
screen "33_Mode_Station_3" 800x480
   Button "Button_5" at 299,208 size 88x48; TextOff 'Stop / AUTO'
      on Press: SetTag("DB_HMI_ARG1_Seq1_Cmd_Auto(2)", 1)
      on Release: SetTag("DB_HMI_ARG1_Seq1_Cmd_Auto(2)", 0)
   Button "Button_6" at 405,208 size 88x48; TextOff 'Reset / MAN'
      on Press: SetTag("DB_HMI_ARG1_Seq1_Cmd_Man(2)", 1)
      on Release: SetTag("DB_HMI_ARG1_Seq1_Cmd_Man(2)", 0)
   Button "Button_1" at 177,283 size 440x40; TextOn 'CLOSE / SCHLIESSEN'; TextOff 'CLOSE / SCHLIESSEN'
      on Click: function_efd93a16()
      Appearance <- "ButtonDown"
   TextField "txtTitleBar" at 16,8 size 495x32; Text 'Operating Mode / Betriebsmodus'
   TextField "txtParameter7_3" at 193,122 size 163x24; Text 'Current Mode / Aktueller Modus'
   TextField "Auto" at 193,149 size 37x20; Text 'Auto'
      Visibility <- "DB_HMI_ARG1_Seq1_Status_Auto(2)"
   TextField "Manual" at 193,148 size 32x20; Text 'Man'
      Visibility <- "DB_HMI_ARG1_Seq1_Status_Man(2)"

screen "34_Mode_Station_4" 800x480
   Button "Button_5" at 299,208 size 88x48; TextOff 'Stop / AUTO'
      on Press: SetTag("DB_HMI_ARG1_Seq1_Cmd_Auto(3)", 1)
      on Release: SetTag("DB_HMI_ARG1_Seq1_Cmd_Auto(3)", 0)
   Button "Button_6" at 405,208 size 88x48; TextOff 'Reset / MAN'
      on Press: SetTag("DB_HMI_ARG1_Seq1_Cmd_Man(3)", 1)
      on Release: SetTag("DB_HMI_ARG1_Seq1_Cmd_Man(3)", 0)
   Button "Button_1" at 177,283 size 440x40; TextOn 'CLOSE / SCHLIESSEN'; TextOff 'CLOSE / SCHLIESSEN'
      on Click: function_efd93a16()
      Appearance <- "ButtonDown"
   TextField "txtTitleBar" at 16,8 size 495x32; Text 'Operating Mode / Betriebsmodus'
   TextField "txtParameter7_3" at 193,122 size 163x24; Text 'Current Mode / Aktueller Modus'
   TextField "Auto" at 193,149 size 37x20; Text 'Auto'
      Visibility <- "DB_HMI_ARG1_Seq1_Status_Auto(3)"
   TextField "Manual" at 193,148 size 32x20; Text 'Man'
      Visibility <- "DB_HMI_ARG1_Seq1_Status_Man(3)"

screen "35_Mode_Station_5" 800x480
   Button "Button_5" at 299,208 size 88x48; TextOff 'Stop / AUTO'
      on Press: SetTag("DB_HMI_ARG1_Seq1_Cmd_Auto(4)", 1)
      on Release: SetTag("DB_HMI_ARG1_Seq1_Cmd_Auto(4)", 0)
   Button "Button_6" at 405,208 size 88x48; TextOff 'Reset / MAN'
      on Press: SetTag("DB_HMI_ARG1_Seq1_Cmd_Man(4)", 1)
      on Release: SetTag("DB_HMI_ARG1_Seq1_Cmd_Man(4)", 0)
   Button "Button_1" at 177,283 size 440x40; TextOn 'CLOSE / SCHLIESSEN'; TextOff 'CLOSE / SCHLIESSEN'
      on Click: function_efd93a16()
      Appearance <- "ButtonDown"
   TextField "txtTitleBar" at 16,8 size 495x32; Text 'Operating Mode / Betriebsmodus'
   TextField "txtParameter7_3" at 193,122 size 163x24; Text 'Current Mode / Aktueller Modus'
   TextField "Auto" at 193,149 size 37x20; Text 'Auto'
      Visibility <- "DB_HMI_ARG1_Seq1_Status_Auto(4)"
   TextField "Manual" at 193,148 size 32x20; Text 'Man'
      Visibility <- "DB_HMI_ARG1_Seq1_Status_Man(4)"

screen "40_SimValues_1" 800x480, template "31_SimValues_1"
   GraphicView "gfxDarkBackground" at 0,0 size 800x480; Picture "PopUpBackground"
      Visibility <- "PopUpBackground"
   TextField "txtParameter1_2" at 246,136 size 42x25; Text 'Step 2 / Parameter 1'
   TextField "txtParameter1_3" at 316,136 size 102x25; Text 'Step 3 / Parameter 1'
   TextField "txtParameter1_4" at 386,136 size 102x25; Text 'Step 4 / Parameter 1'
   TextField "txtParameter1_5" at 456,136 size 102x25; Text 'Step 5 / Parameter 1'
   TextField "txtParameter1_6" at 526,136 size 102x25; Text 'Step 6 / Parameter 1'
   TextField "txtParameter1_8" at 596,136 size 102x25; Text 'Step 7 / Parameter 1'
   TextField "txtParameter1_9" at 666,136 size 102x25; Text 'Step 8 / Parameter 1'
   TextField "txtParameter1_10" at 176,136 size 45x25; Text 'Step 1 / Parameter 1'
   TextField "txtParameter1_11" at 736,136 size 46x25; Text 'Step 9 / Parameter 1'
   TextField "txtParameter1_1" at 104,136 size 45x25; Text 'Branch / Parameter 1'
   TextField "txtParameter1_7" at 32,136 size 45x25; Text 'Car / Parameter 1'
   GraphicView "Graphic view_1" at 33,184 size 40x40; Picture "Car_Red"
   GraphicView "Graphic view_3" at 33,249 size 40x40; Picture "Car_Green"
   GraphicView "Graphic view_4" at 33,308 size 40x40; Picture "Car_Blue_1"
   TextField "Text field_3" at 121,191 size 15x23; Text '1'
      Visibility <- "InScreenTabState"
   TextField "Text field_1" at 121,256 size 15x23; Text '2'
      Visibility <- "InScreenTabState"
   TextField "Text field_2" at 121,321 size 15x23; Text '2'
      Visibility <- "InScreenTabState"
   Button "Button_1" at 176,186 size 38x32; TextOff 'Text'
      on Click: SetTag("DB_HMI_ARG1_Seq1_DelaySelect_Red{2}", 1)
   Button "Button_2" at 245,186 size 38x32; TextOff 'Text'
      on Click: SetTag("DB_HMI_ARG1_Seq1_DelaySelect_Red{3}", 1)
   Button "Button_3" at 315,186 size 38x32; TextOff 'Text'
      on Click: SetTag("DB_HMI_ARG1_Seq1_DelaySelect_Red{4}", 1)
   Button "Button_4" at 385,186 size 38x32; TextOff 'Text'
      on Click: SetTag("DB_HMI_ARG1_Seq1_DelaySelect_Red{5}", 1)
   Button "Button_5" at 455,186 size 38x32; TextOff 'Text'
      on Click: SetTag("DB_HMI_ARG1_Seq1_DelaySelect_Red{6}", 1)
   Button "Button_6" at 525,186 size 38x32; TextOff 'Text'
      on Click: SetTag("DB_HMI_ARG1_Seq1_DelaySelect_Red{7}", 1)
   Button "Button_8" at 595,186 size 38x32; TextOff 'Text'
      on Click: SetTag("DB_HMI_ARG1_Seq1_DelaySelect_Red{8}", 1)
   Button "Button_9" at 665,186 size 38x32; TextOff 'Text'
      on Click: SetTag("DB_HMI_ARG1_Seq1_DelaySelect_Red{9}", 1)
   Button "Button_10" at 735,186 size 38x32; TextOff 'Text'
      on Click: SetTag("DB_HMI_ARG1_Seq1_DelaySelect_Red{10}", 1)
   Button "Button_17" at 176,250 size 38x32; TextOff 'Text'
      on Click: SetTag("DB_HMI_ARG1_Seq1_DelaySelect_Green{2}", 1)
   Button "Button_7" at 246,250 size 38x32; TextOff 'Text'
      on Click: SetTag("DB_HMI_ARG1_Seq1_DelaySelect_Green{3}", 1)
   Button "Button_11" at 316,250 size 38x32; TextOff 'Text'
      on Click: SetTag("DB_HMI_ARG1_Seq1_DelaySelect_Green{4}", 1)
   Button "Button_12" at 386,250 size 38x32; TextOff 'Text'
      on Click: SetTag("DB_HMI_ARG1_Seq1_DelaySelect_Green{5}", 1)
   Button "Button_13" at 456,250 size 38x32; TextOff 'Text'
      on Click: SetTag("DB_HMI_ARG1_Seq1_DelaySelect_Green{6}", 1)
   Button "Button_14" at 526,250 size 38x32; TextOff 'Text'
      on Click: SetTag("DB_HMI_ARG1_Seq1_DelaySelect_Green{7}", 1)
   Button "Button_15" at 596,250 size 38x32; TextOff 'Text'
      on Click: SetTag("DB_HMI_ARG1_Seq1_DelaySelect_Green{8}", 1)
   Button "Button_16" at 666,250 size 38x32; TextOff 'Text'
      on Click: SetTag("DB_HMI_ARG1_Seq1_DelaySelect_Green{9}", 1)
   Button "Button_18" at 736,250 size 38x32; TextOff 'Text'
      on Click: SetTag("DB_HMI_ARG1_Seq1_DelaySelect_Green{10}", 1)
   Button "Button_26" at 176,314 size 38x32; TextOff 'Text'
      on Click: SetTag("DB_HMI_ARG1_Seq1_DelaySelect_Blue{2}", 1)
   Button "Button_19" at 246,314 size 38x32; TextOff 'Text'
      on Click: SetTag("DB_HMI_ARG1_Seq1_DelaySelect_Blue{3}", 1)
   Button "Button_20" at 316,314 size 38x32; TextOff 'Text'
      on Click: SetTag("DB_HMI_ARG1_Seq1_DelaySelect_Blue{4}", 1)
   Button "Button_21" at 386,314 size 38x32; TextOff 'Text'
      on Click: SetTag("DB_HMI_ARG1_Seq1_DelaySelect_Blue{5}", 1)
   Button "Button_22" at 456,314 size 38x32; TextOff 'Text'
      on Click: SetTag("DB_HMI_ARG1_Seq1_DelaySelect_Blue{6}", 1)
   Button "Button_23" at 526,314 size 38x32; TextOff 'Text'
      on Click: SetTag("DB_HMI_ARG1_Seq1_DelaySelect_Blue{7}", 1)
   Button "Button_24" at 596,314 size 38x32; TextOff 'Text'
      on Click: SetTag("DB_HMI_ARG1_Seq1_DelaySelect_Blue{8}", 1)
   Button "Button_25" at 666,314 size 38x32; TextOff 'Text'
      on Click: SetTag("DB_HMI_ARG1_Seq1_DelaySelect_Blue{9}", 1)
   Button "Button_27" at 736,314 size 38x32; TextOff 'Text'
      on Click: SetTag("DB_HMI_ARG1_Seq1_DelaySelect_Blue{10}", 1)
   Button "Button_28" at 176,186 size 38x32; TextOff 'Text'
      on Click: SetTag("DB_HMI_ARG1_Seq1_DelaySelect_Red{2}", 0)
      Visibility <- "DB_HMI_ARG1_Seq1_DelaySelect_Red{2}"
   Button "Button_29" at 245,186 size 38x32; TextOff 'Text'
      on Click: SetTag("DB_HMI_ARG1_Seq1_DelaySelect_Red{3}", 0)
      Visibility <- "DB_HMI_ARG1_Seq1_DelaySelect_Red{3}"
   Button "Button_30" at 315,186 size 38x32; TextOff 'Text'
      on Click: SetTag("DB_HMI_ARG1_Seq1_DelaySelect_Red{4}", 0)
      Visibility <- "DB_HMI_ARG1_Seq1_DelaySelect_Red{4}"
   Button "Button_31" at 385,186 size 38x32; TextOff 'Text'
      on Click: SetTag("DB_HMI_ARG1_Seq1_DelaySelect_Red{5}", 0)
      Visibility <- "DB_HMI_ARG1_Seq1_DelaySelect_Red{5}"
   Button "Button_32" at 455,186 size 38x32; TextOff 'Text'
      on Click: SetTag("DB_HMI_ARG1_Seq1_DelaySelect_Red{6}", 0)
      Visibility <- "DB_HMI_ARG1_Seq1_DelaySelect_Red{6}"
   Button "Button_33" at 525,186 size 38x32; TextOff 'Text'
      on Click: SetTag("DB_HMI_ARG1_Seq1_DelaySelect_Red{7}", 0)
      Visibility <- "DB_HMI_ARG1_Seq1_DelaySelect_Red{7}"
   Button "Button_34" at 595,186 size 38x32; TextOff 'Text'
      on Click: SetTag("DB_HMI_ARG1_Seq1_DelaySelect_Red{8}", 0)
      Visibility <- "DB_HMI_ARG1_Seq1_DelaySelect_Red{8}"
   Button "Button_35" at 665,186 size 38x32; TextOff 'Text'
      on Click: SetTag("DB_HMI_ARG1_Seq1_DelaySelect_Red{9}", 0)
      Visibility <- "DB_HMI_ARG1_Seq1_DelaySelect_Red{9}"
   Button "Button_36" at 735,186 size 38x32; TextOff 'Text'
      on Click: SetTag("DB_HMI_ARG1_Seq1_DelaySelect_Red{10}", 0)
      Visibility <- "DB_HMI_ARG1_Seq1_DelaySelect_Red{10}"
   Button "Button_37" at 176,250 size 38x32; TextOff 'Text'
      on Click: SetTag("DB_HMI_ARG1_Seq1_DelaySelect_Green{2}", 0)
      Visibility <- "DB_HMI_ARG1_Seq1_DelaySelect_Green{2}"
   Button "Button_38" at 246,250 size 38x32; TextOff 'Text'
      on Click: SetTag("DB_HMI_ARG1_Seq1_DelaySelect_Green{3}", 0)
      Visibility <- "DB_HMI_ARG1_Seq1_DelaySelect_Green{3}"
   Button "Button_39" at 316,250 size 38x32; TextOff 'Text'
      on Click: SetTag("DB_HMI_ARG1_Seq1_DelaySelect_Green{4}", 0)
      Visibility <- "DB_HMI_ARG1_Seq1_DelaySelect_Green{4}"
   Button "Button_40" at 386,250 size 38x32; TextOff 'Text'
      on Click: SetTag("DB_HMI_ARG1_Seq1_DelaySelect_Green{5}", 0)
      Visibility <- "DB_HMI_ARG1_Seq1_DelaySelect_Green{5}"
   Button "Button_41" at 456,250 size 38x32; TextOff 'Text'
      on Click: SetTag("DB_HMI_ARG1_Seq1_DelaySelect_Green{6}", 0)
      Visibility <- "DB_HMI_ARG1_Seq1_DelaySelect_Green{6}"
   Button "Button_42" at 526,250 size 38x32; TextOff 'Text'
      on Click: SetTag("DB_HMI_ARG1_Seq1_DelaySelect_Green{7}", 0)
      Visibility <- "DB_HMI_ARG1_Seq1_DelaySelect_Green{7}"
   Button "Button_43" at 596,250 size 38x32; TextOff 'Text'
      on Click: SetTag("DB_HMI_ARG1_Seq1_DelaySelect_Green{8}", 0)
      Visibility <- "DB_HMI_ARG1_Seq1_DelaySelect_Green{8}"
   Button "Button_44" at 666,250 size 38x32; TextOff 'Text'
      on Click: SetTag("DB_HMI_ARG1_Seq1_DelaySelect_Green{9}", 0)
      Visibility <- "DB_HMI_ARG1_Seq1_DelaySelect_Green{9}"
   Button "Button_45" at 736,250 size 38x32; TextOff 'Text'
      on Click: SetTag("DB_HMI_ARG1_Seq1_DelaySelect_Green{10}", 0)
      Visibility <- "DB_HMI_ARG1_Seq1_DelaySelect_Green{10}"
   Button "Button_46" at 176,314 size 38x32; TextOff 'Text'
      on Click: SetTag("DB_HMI_ARG1_Seq1_DelaySelect_Blue{2}", 0)
      Visibility <- "DB_HMI_ARG1_Seq1_DelaySelect_Blue{2}"
   Button "Button_47" at 246,314 size 38x32; TextOff 'Text'
      on Click: SetTag("DB_HMI_ARG1_Seq1_DelaySelect_Blue{3}", 0)
      Visibility <- "DB_HMI_ARG1_Seq1_DelaySelect_Blue{3}"
   Button "Button_48" at 316,314 size 38x32; TextOff 'Text'
      on Click: SetTag("DB_HMI_ARG1_Seq1_DelaySelect_Blue{4}", 0)
      Visibility <- "DB_HMI_ARG1_Seq1_DelaySelect_Blue{4}"
   Button "Button_49" at 386,314 size 38x32; TextOff 'Text'
      on Click: SetTag("DB_HMI_ARG1_Seq1_DelaySelect_Blue{5}", 0)
      Visibility <- "DB_HMI_ARG1_Seq1_DelaySelect_Blue{5}"
   Button "Button_50" at 456,314 size 38x32; TextOff 'Text'
      on Click: SetTag("DB_HMI_ARG1_Seq1_DelaySelect_Blue{6}", 0)
      Visibility <- "DB_HMI_ARG1_Seq1_DelaySelect_Blue{6}"
   Button "Button_51" at 526,314 size 38x32; TextOff 'Text'
      on Click: SetTag("DB_HMI_ARG1_Seq1_DelaySelect_Blue{7}", 0)
      Visibility <- "DB_HMI_ARG1_Seq1_DelaySelect_Blue{7}"
   Button "Button_52" at 596,314 size 38x32; TextOff 'Text'
      on Click: SetTag("DB_HMI_ARG1_Seq1_DelaySelect_Blue{8}", 0)
      Visibility <- "DB_HMI_ARG1_Seq1_DelaySelect_Blue{8}"
   Button "Button_53" at 666,314 size 38x32; TextOff 'Text'
      on Click: SetTag("DB_HMI_ARG1_Seq1_DelaySelect_Blue{9}", 0)
      Visibility <- "DB_HMI_ARG1_Seq1_DelaySelect_Blue{9}"
   Button "Button_54" at 736,314 size 38x32; TextOff 'Text'
      on Click: SetTag("DB_HMI_ARG1_Seq1_DelaySelect_Blue{10}", 0)
      Visibility <- "DB_HMI_ARG1_Seq1_DelaySelect_Blue{10}"
   Button "Button_55" at 619,378 size 165x40; TextOff 'Reset / Alle Quittieren'; PictureOff "More_Icon"
      on ReleaseLeft: ResetBit("Ext_AckSafety_DB_ack")
      on Press: SetTag("DB_HMI_ARG1_Seq1_Cmd_DelayReset", 1)
      on PressLeft: SetBit("Ext_AckSafety_DB_ack")
      on Release: SetTag("DB_HMI_ARG1_Seq1_Cmd_DelayReset", 0)
      ObjectEnable <- "DB_HMI_ARG1_Seq1_Cmd_DelayReset"

screen "40_SimValues_2" 800x480, template "31_SimValues_1"
   GraphicView "gfxDarkBackground" at 0,0 size 800x480; Picture "PopUpBackground"
      Visibility <- "PopUpBackground"
   TextField "txtParameter1_2" at 246,136 size 42x25; Text 'Step 2 / Parameter 1'
   TextField "txtParameter1_3" at 316,136 size 102x25; Text 'Step 3 / Parameter 1'
   TextField "txtParameter1_4" at 386,136 size 102x25; Text 'Step 4 / Parameter 1'
   TextField "txtParameter1_5" at 456,136 size 102x25; Text 'Step 5 / Parameter 1'
   TextField "txtParameter1_6" at 526,136 size 102x25; Text 'Step 6 / Parameter 1'
   TextField "txtParameter1_8" at 596,136 size 102x25; Text 'Step 7 / Parameter 1'
   TextField "txtParameter1_9" at 666,136 size 102x25; Text 'Step 8 / Parameter 1'
   TextField "txtParameter1_10" at 176,136 size 45x25; Text 'Step 1 / Parameter 1'
   TextField "txtParameter1_11" at 736,136 size 46x25; Text 'Step 9 / Parameter 1'
   TextField "txtParameter1_1" at 104,136 size 45x25; Text 'Branch / Parameter 1'
   TextField "txtParameter1_7" at 32,136 size 45x25; Text 'Car / Parameter 1'
   GraphicView "Graphic view_1" at 33,184 size 40x40; Picture "Car_Red"
   GraphicView "Graphic view_3" at 33,249 size 40x40; Picture "Car_Green"
   GraphicView "Graphic view_4" at 33,308 size 40x40; Picture "Car_Blue_1"
   TextField "Text field_3" at 121,191 size 15x23; Text '1'
      Visibility <- "InScreenTabState"
   TextField "Text field_1" at 121,256 size 15x23; Text '2'
      Visibility <- "InScreenTabState"
   TextField "Text field_2" at 121,321 size 15x23; Text '2'
      Visibility <- "InScreenTabState"
   Button "Button_1" at 176,186 size 38x32; TextOff 'Text'
      on Click: SetTag("DB_HMI_ARG1_Seq1_DelaySelect_Red{2}(1)", 1)
   Button "Button_2" at 245,186 size 38x32; TextOff 'Text'
      on Click: SetTag("DB_HMI_ARG1_Seq1_DelaySelect_Red{3}(1)", 1)
   Button "Button_3" at 315,186 size 38x32; TextOff 'Text'
      on Click: SetTag("DB_HMI_ARG1_Seq1_DelaySelect_Red{4}(1)", 1)
   Button "Button_4" at 385,186 size 38x32; TextOff 'Text'
      on Click: SetTag("DB_HMI_ARG1_Seq1_DelaySelect_Red{5}(1)", 1)
   Button "Button_5" at 455,186 size 38x32; TextOff 'Text'
      on Click: SetTag("DB_HMI_ARG1_Seq1_DelaySelect_Red{6}(1)", 1)
   Button "Button_6" at 525,186 size 38x32; TextOff 'Text'
      on Click: SetTag("DB_HMI_ARG1_Seq1_DelaySelect_Red{7}(1)", 1)
   Button "Button_8" at 595,186 size 38x32; TextOff 'Text'
      on Click: SetTag("DB_HMI_ARG1_Seq1_DelaySelect_Red{8}(1)", 1)
   Button "Button_9" at 665,186 size 38x32; TextOff 'Text'
      on Click: SetTag("DB_HMI_ARG1_Seq1_DelaySelect_Red{9}(1)", 1)
   Button "Button_10" at 735,186 size 38x32; TextOff 'Text'
      on Click: SetTag("DB_HMI_ARG1_Seq1_DelaySelect_Red{10}(1)", 1)
   Button "Button_17" at 176,250 size 38x32; TextOff 'Text'
      on Click: SetTag("DB_HMI_ARG1_Seq1_DelaySelect_Green{2}(1)", 1)
   Button "Button_7" at 246,250 size 38x32; TextOff 'Text'
      on Click: SetTag("DB_HMI_ARG1_Seq1_DelaySelect_Green{3}(1)", 1)
   Button "Button_11" at 316,250 size 38x32; TextOff 'Text'
      on Click: SetTag("DB_HMI_ARG1_Seq1_DelaySelect_Green{4}(1)", 1)
   Button "Button_12" at 386,250 size 38x32; TextOff 'Text'
      on Click: SetTag("DB_HMI_ARG1_Seq1_DelaySelect_Green{5}(1)", 1)
   Button "Button_13" at 456,250 size 38x32; TextOff 'Text'
      on Click: SetTag("DB_HMI_ARG1_Seq1_DelaySelect_Green{6}(1)", 1)
   Button "Button_14" at 526,250 size 38x32; TextOff 'Text'
      on Click: SetTag("DB_HMI_ARG1_Seq1_DelaySelect_Green{7}(1)", 1)
   Button "Button_15" at 596,250 size 38x32; TextOff 'Text'
      on Click: SetTag("DB_HMI_ARG1_Seq1_DelaySelect_Green{8}(1)", 1)
   Button "Button_16" at 666,250 size 38x32; TextOff 'Text'
      on Click: SetTag("DB_HMI_ARG1_Seq1_DelaySelect_Green{9}(1)", 1)
   Button "Button_18" at 736,250 size 38x32; TextOff 'Text'
      on Click: SetTag("DB_HMI_ARG1_Seq1_DelaySelect_Green{10}(1)", 1)
   Button "Button_26" at 176,314 size 38x32; TextOff 'Text'
      on Click: SetTag("DB_HMI_ARG1_Seq1_DelaySelect_Blue{2}(1)", 1)
   Button "Button_19" at 246,314 size 38x32; TextOff 'Text'
      on Click: SetTag("DB_HMI_ARG1_Seq1_DelaySelect_Blue{3}(1)", 1)
   Button "Button_20" at 316,314 size 38x32; TextOff 'Text'
      on Click: SetTag("DB_HMI_ARG1_Seq1_DelaySelect_Blue{4}(1)", 1)
   Button "Button_21" at 386,314 size 38x32; TextOff 'Text'
      on Click: SetTag("DB_HMI_ARG1_Seq1_DelaySelect_Blue{5}(1)", 1)
   Button "Button_22" at 456,314 size 38x32; TextOff 'Text'
      on Click: SetTag("DB_HMI_ARG1_Seq1_DelaySelect_Blue{6}(1)", 1)
   Button "Button_23" at 526,314 size 38x32; TextOff 'Text'
      on Click: SetTag("DB_HMI_ARG1_Seq1_DelaySelect_Blue{7}(1)", 1)
   Button "Button_24" at 596,314 size 38x32; TextOff 'Text'
      on Click: SetTag("DB_HMI_ARG1_Seq1_DelaySelect_Blue{8}(1)", 1)
   Button "Button_25" at 666,314 size 38x32; TextOff 'Text'
      on Click: SetTag("DB_HMI_ARG1_Seq1_DelaySelect_Blue{9}(1)", 1)
   Button "Button_27" at 736,314 size 38x32; TextOff 'Text'
      on Click: SetTag("DB_HMI_ARG1_Seq1_DelaySelect_Blue{10}(1)", 1)
   Button "Button_28" at 176,186 size 38x32; TextOff 'Text'
      on Click: SetTag("DB_HMI_ARG1_Seq1_DelaySelect_Red{2}(1)", 0)
      Visibility <- "DB_HMI_ARG1_Seq1_DelaySelect_Red{2}(1)"
   Button "Button_29" at 245,186 size 38x32; TextOff 'Text'
      on Click: SetTag("DB_HMI_ARG1_Seq1_DelaySelect_Red{3}(1)", 0)
      Visibility <- "DB_HMI_ARG1_Seq1_DelaySelect_Red{3}(1)"
   Button "Button_30" at 315,186 size 38x32; TextOff 'Text'
      on Click: SetTag("DB_HMI_ARG1_Seq1_DelaySelect_Red{4}(1)", 0)
      Visibility <- "DB_HMI_ARG1_Seq1_DelaySelect_Red{4}(1)"
   Button "Button_31" at 385,186 size 38x32; TextOff 'Text'
      on Click: SetTag("DB_HMI_ARG1_Seq1_DelaySelect_Red{5}(1)", 0)
      Visibility <- "DB_HMI_ARG1_Seq1_DelaySelect_Red{5}(1)"
   Button "Button_32" at 455,186 size 38x32; TextOff 'Text'
      on Click: SetTag("DB_HMI_ARG1_Seq1_DelaySelect_Red{6}(1)", 0)
      Visibility <- "DB_HMI_ARG1_Seq1_DelaySelect_Red{6}(1)"
   Button "Button_33" at 525,186 size 38x32; TextOff 'Text'
      on Click: SetTag("DB_HMI_ARG1_Seq1_DelaySelect_Red{7}(1)", 0)
      Visibility <- "DB_HMI_ARG1_Seq1_DelaySelect_Red{7}(1)"
   Button "Button_34" at 595,186 size 38x32; TextOff 'Text'
      on Click: SetTag("DB_HMI_ARG1_Seq1_DelaySelect_Red{8}(1)", 0)
      Visibility <- "DB_HMI_ARG1_Seq1_DelaySelect_Red{8}(1)"
   Button "Button_35" at 665,186 size 38x32; TextOff 'Text'
      on Click: SetTag("DB_HMI_ARG1_Seq1_DelaySelect_Red{9}(1)", 0)
      Visibility <- "DB_HMI_ARG1_Seq1_DelaySelect_Red{9}(1)"
   Button "Button_36" at 735,186 size 38x32; TextOff 'Text'
      on Click: SetTag("DB_HMI_ARG1_Seq1_DelaySelect_Red{10}(1)", 0)
      Visibility <- "DB_HMI_ARG1_Seq1_DelaySelect_Red{10}(1)"
   Button "Button_37" at 176,250 size 38x32; TextOff 'Text'
      on Click: SetTag("DB_HMI_ARG1_Seq1_DelaySelect_Green{2}(1)", 0)
      Visibility <- "DB_HMI_ARG1_Seq1_DelaySelect_Green{2}(1)"
   Button "Button_38" at 246,250 size 38x32; TextOff 'Text'
      on Click: SetTag("DB_HMI_ARG1_Seq1_DelaySelect_Green{3}(1)", 0)
      Visibility <- "DB_HMI_ARG1_Seq1_DelaySelect_Green{3}(1)"
   Button "Button_39" at 316,250 size 38x32; TextOff 'Text'
      on Click: SetTag("DB_HMI_ARG1_Seq1_DelaySelect_Green{4}(1)", 0)
      Visibility <- "DB_HMI_ARG1_Seq1_DelaySelect_Green{4}(1)"
   Button "Button_40" at 386,250 size 38x32; TextOff 'Text'
      on Click: SetTag("DB_HMI_ARG1_Seq1_DelaySelect_Green{5}(1)", 0)
      Visibility <- "DB_HMI_ARG1_Seq1_DelaySelect_Green{5}(1)"
   Button "Button_41" at 456,250 size 38x32; TextOff 'Text'
      on Click: SetTag("DB_HMI_ARG1_Seq1_DelaySelect_Green{6}(1)", 0)
      Visibility <- "DB_HMI_ARG1_Seq1_DelaySelect_Green{6}(1)"
   Button "Button_42" at 526,250 size 38x32; TextOff 'Text'
      on Click: SetTag("DB_HMI_ARG1_Seq1_DelaySelect_Green{7}(1)", 0)
      Visibility <- "DB_HMI_ARG1_Seq1_DelaySelect_Green{7}(1)"
   Button "Button_43" at 596,250 size 38x32; TextOff 'Text'
      on Click: SetTag("DB_HMI_ARG1_Seq1_DelaySelect_Green{8}(1)", 0)
      Visibility <- "DB_HMI_ARG1_Seq1_DelaySelect_Green{8}(1)"
   Button "Button_44" at 666,250 size 38x32; TextOff 'Text'
      on Click: SetTag("DB_HMI_ARG1_Seq1_DelaySelect_Green{9}(1)", 0)
      Visibility <- "DB_HMI_ARG1_Seq1_DelaySelect_Green{9}(1)"
   Button "Button_45" at 736,250 size 38x32; TextOff 'Text'
      on Click: SetTag("DB_HMI_ARG1_Seq1_DelaySelect_Green{10}(1)", 0)
      Visibility <- "DB_HMI_ARG1_Seq1_DelaySelect_Green{10}(1)"
   Button "Button_46" at 176,314 size 38x32; TextOff 'Text'
      on Click: SetTag("DB_HMI_ARG1_Seq1_DelaySelect_Blue{2}(1)", 0)
      Visibility <- "DB_HMI_ARG1_Seq1_DelaySelect_Blue{2}(1)"
   Button "Button_47" at 246,314 size 38x32; TextOff 'Text'
      on Click: SetTag("DB_HMI_ARG1_Seq1_DelaySelect_Blue{3}(1)", 0)
      Visibility <- "DB_HMI_ARG1_Seq1_DelaySelect_Blue{3}(1)"
   Button "Button_48" at 316,314 size 38x32; TextOff 'Text'
      on Click: SetTag("DB_HMI_ARG1_Seq1_DelaySelect_Blue{4}(1)", 0)
      Visibility <- "DB_HMI_ARG1_Seq1_DelaySelect_Blue{4}(1)"
   Button "Button_49" at 386,314 size 38x32; TextOff 'Text'
      on Click: SetTag("DB_HMI_ARG1_Seq1_DelaySelect_Blue{5}(1)", 0)
      Visibility <- "DB_HMI_ARG1_Seq1_DelaySelect_Blue{5}(1)"
   Button "Button_50" at 456,314 size 38x32; TextOff 'Text'
      on Click: SetTag("DB_HMI_ARG1_Seq1_DelaySelect_Blue{6}(1)", 0)
      Visibility <- "DB_HMI_ARG1_Seq1_DelaySelect_Blue{6}(1)"
   Button "Button_51" at 526,314 size 38x32; TextOff 'Text'
      on Click: SetTag("DB_HMI_ARG1_Seq1_DelaySelect_Blue{7}(1)", 0)
      Visibility <- "DB_HMI_ARG1_Seq1_DelaySelect_Blue{7}(1)"
   Button "Button_52" at 596,314 size 38x32; TextOff 'Text'
      on Click: SetTag("DB_HMI_ARG1_Seq1_DelaySelect_Blue{8}(1)", 0)
      Visibility <- "DB_HMI_ARG1_Seq1_DelaySelect_Blue{8}(1)"
   Button "Button_53" at 666,314 size 38x32; TextOff 'Text'
      on Click: SetTag("DB_HMI_ARG1_Seq1_DelaySelect_Blue{9}(1)", 0)
      Visibility <- "DB_HMI_ARG1_Seq1_DelaySelect_Blue{9}(1)"
   Button "Button_54" at 736,314 size 38x32; TextOff 'Text'
      on Click: SetTag("DB_HMI_ARG1_Seq1_DelaySelect_Blue{10}(1)", 0)
      Visibility <- "DB_HMI_ARG1_Seq1_DelaySelect_Blue{10}(1)"
   Button "Button_55" at 619,378 size 165x40; TextOff 'Reset / Alle Quittieren'; PictureOff "More_Icon"
      on ReleaseLeft: ResetBit("Ext_AckSafety_DB_ack")
      on PressLeft: SetBit("Ext_AckSafety_DB_ack")
      on Release: SetTag("DB_HMI_ARG1_Seq1_Cmd_DelayReset(1)", 0)
      on Press: SetTag("DB_HMI_ARG1_Seq1_Cmd_DelayReset(1)", 1)
      ObjectEnable <- "DB_HMI_ARG1_Seq1_Cmd_DelayReset"

screen "40_SimValues_3" 800x480, template "31_SimValues_1"
   GraphicView "gfxDarkBackground" at 0,0 size 800x480; Picture "PopUpBackground"
      Visibility <- "PopUpBackground"
   TextField "txtParameter1_2" at 246,136 size 42x25; Text 'Step 2 / Parameter 1'
   TextField "txtParameter1_3" at 316,136 size 102x25; Text 'Step 3 / Parameter 1'
   TextField "txtParameter1_4" at 386,136 size 102x25; Text 'Step 4 / Parameter 1'
   TextField "txtParameter1_5" at 456,136 size 102x25; Text 'Step 5 / Parameter 1'
   TextField "txtParameter1_6" at 526,136 size 102x25; Text 'Step 6 / Parameter 1'
   TextField "txtParameter1_8" at 596,136 size 102x25; Text 'Step 7 / Parameter 1'
   TextField "txtParameter1_9" at 666,136 size 102x25; Text 'Step 8 / Parameter 1'
   TextField "txtParameter1_10" at 176,136 size 45x25; Text 'Step 1 / Parameter 1'
   TextField "txtParameter1_11" at 736,136 size 46x25; Text 'Step 9 / Parameter 1'
   TextField "txtParameter1_1" at 104,136 size 45x25; Text 'Branch / Parameter 1'
   TextField "txtParameter1_7" at 32,136 size 45x25; Text 'Car / Parameter 1'
   GraphicView "Graphic view_1" at 33,184 size 40x40; Picture "Car_Red"
   GraphicView "Graphic view_3" at 33,249 size 40x40; Picture "Car_Green"
   GraphicView "Graphic view_4" at 33,308 size 40x40; Picture "Car_Blue_1"
   TextField "Text field_3" at 121,191 size 15x23; Text '1'
      Visibility <- "InScreenTabState"
   TextField "Text field_1" at 121,256 size 15x23; Text '2'
      Visibility <- "InScreenTabState"
   TextField "Text field_2" at 121,321 size 15x23; Text '2'
      Visibility <- "InScreenTabState"
   Button "Button_1" at 176,186 size 38x32; TextOff 'Text'
      on Click: SetTag("DB_HMI_ARG1_Seq1_DelaySelect_Red{2}(2)", 1)
   Button "Button_2" at 245,186 size 38x32; TextOff 'Text'
      on Click: SetTag("DB_HMI_ARG1_Seq1_DelaySelect_Red{3}(2)", 1)
   Button "Button_3" at 315,186 size 38x32; TextOff 'Text'
      on Click: SetTag("DB_HMI_ARG1_Seq1_DelaySelect_Red{4}(2)", 1)
   Button "Button_4" at 385,186 size 38x32; TextOff 'Text'
      on Click: SetTag("DB_HMI_ARG1_Seq1_DelaySelect_Red{5}(2)", 1)
   Button "Button_5" at 455,186 size 38x32; TextOff 'Text'
      on Click: SetTag("DB_HMI_ARG1_Seq1_DelaySelect_Red{6}(2)", 1)
   Button "Button_6" at 525,186 size 38x32; TextOff 'Text'
      on Click: SetTag("DB_HMI_ARG1_Seq1_DelaySelect_Red{7}(2)", 1)
   Button "Button_8" at 595,186 size 38x32; TextOff 'Text'
      on Click: SetTag("DB_HMI_ARG1_Seq1_DelaySelect_Red{8}(2)", 1)
   Button "Button_9" at 665,186 size 38x32; TextOff 'Text'
      on Click: SetTag("DB_HMI_ARG1_Seq1_DelaySelect_Red{9}(2)", 1)
   Button "Button_10" at 735,186 size 38x32; TextOff 'Text'
      on Click: SetTag("DB_HMI_ARG1_Seq1_DelaySelect_Red{10}(2)", 1)
   Button "Button_17" at 176,250 size 38x32; TextOff 'Text'
      on Click: SetTag("DB_HMI_ARG1_Seq1_DelaySelect_Green{2}(2)", 1)
   Button "Button_7" at 246,250 size 38x32; TextOff 'Text'
      on Click: SetTag("DB_HMI_ARG1_Seq1_DelaySelect_Green{3}(2)", 1)
   Button "Button_11" at 316,250 size 38x32; TextOff 'Text'
      on Click: SetTag("DB_HMI_ARG1_Seq1_DelaySelect_Green{4}(2)", 1)
   Button "Button_12" at 386,250 size 38x32; TextOff 'Text'
      on Click: SetTag("DB_HMI_ARG1_Seq1_DelaySelect_Green{5}(2)", 1)
   Button "Button_13" at 456,250 size 38x32; TextOff 'Text'
      on Click: SetTag("DB_HMI_ARG1_Seq1_DelaySelect_Green{6}(2)", 1)
   Button "Button_14" at 526,250 size 38x32; TextOff 'Text'
      on Click: SetTag("DB_HMI_ARG1_Seq1_DelaySelect_Green{7}(2)", 1)
   Button "Button_15" at 596,250 size 38x32; TextOff 'Text'
      on Click: SetTag("DB_HMI_ARG1_Seq1_DelaySelect_Green{8}(2)", 1)
   Button "Button_16" at 666,250 size 38x32; TextOff 'Text'
      on Click: SetTag("DB_HMI_ARG1_Seq1_DelaySelect_Green{9}(2)", 1)
   Button "Button_18" at 736,250 size 38x32; TextOff 'Text'
      on Click: SetTag("DB_HMI_ARG1_Seq1_DelaySelect_Green{10}(2)", 1)
   Button "Button_26" at 176,314 size 38x32; TextOff 'Text'
      on Click: SetTag("DB_HMI_ARG1_Seq1_DelaySelect_Blue{2}(2)", 1)
   Button "Button_19" at 246,314 size 38x32; TextOff 'Text'
      on Click: SetTag("DB_HMI_ARG1_Seq1_DelaySelect_Blue{3}(2)", 1)
   Button "Button_20" at 316,314 size 38x32; TextOff 'Text'
      on Click: SetTag("DB_HMI_ARG1_Seq1_DelaySelect_Blue{4}(2)", 1)
   Button "Button_21" at 386,314 size 38x32; TextOff 'Text'
      on Click: SetTag("DB_HMI_ARG1_Seq1_DelaySelect_Blue{5}(2)", 1)
   Button "Button_22" at 456,314 size 38x32; TextOff 'Text'
      on Click: SetTag("DB_HMI_ARG1_Seq1_DelaySelect_Blue{6}(2)", 1)
   Button "Button_23" at 526,314 size 38x32; TextOff 'Text'
      on Click: SetTag("DB_HMI_ARG1_Seq1_DelaySelect_Blue{7}(2)", 1)
   Button "Button_24" at 596,314 size 38x32; TextOff 'Text'
      on Click: SetTag("DB_HMI_ARG1_Seq1_DelaySelect_Blue{8}(2)", 1)
   Button "Button_25" at 666,314 size 38x32; TextOff 'Text'
      on Click: SetTag("DB_HMI_ARG1_Seq1_DelaySelect_Blue{9}(2)", 1)
   Button "Button_27" at 736,314 size 38x32; TextOff 'Text'
      on Click: SetTag("DB_HMI_ARG1_Seq1_DelaySelect_Blue{10}(2)", 1)
   Button "Button_28" at 176,186 size 38x32; TextOff 'Text'
      on Click: SetTag("DB_HMI_ARG1_Seq1_DelaySelect_Red{2}(2)", 0)
      Visibility <- "DB_HMI_ARG1_Seq1_DelaySelect_Red{2}(2)"
   Button "Button_29" at 245,186 size 38x32; TextOff 'Text'
      on Click: SetTag("DB_HMI_ARG1_Seq1_DelaySelect_Red{3}(2)", 0)
      Visibility <- "DB_HMI_ARG1_Seq1_DelaySelect_Red{3}(2)"
   Button "Button_30" at 315,186 size 38x32; TextOff 'Text'
      on Click: SetTag("DB_HMI_ARG1_Seq1_DelaySelect_Red{4}(2)", 0)
      Visibility <- "DB_HMI_ARG1_Seq1_DelaySelect_Red{4}(2)"
   Button "Button_31" at 385,186 size 38x32; TextOff 'Text'
      on Click: SetTag("DB_HMI_ARG1_Seq1_DelaySelect_Red{5}(2)", 0)
      Visibility <- "DB_HMI_ARG1_Seq1_DelaySelect_Red{5}(2)"
   Button "Button_32" at 455,186 size 38x32; TextOff 'Text'
      on Click: SetTag("DB_HMI_ARG1_Seq1_DelaySelect_Red{6}(2)", 0)
      Visibility <- "DB_HMI_ARG1_Seq1_DelaySelect_Red{6}(2)"
   Button "Button_33" at 525,186 size 38x32; TextOff 'Text'
      on Click: SetTag("DB_HMI_ARG1_Seq1_DelaySelect_Red{7}(2)", 0)
      Visibility <- "DB_HMI_ARG1_Seq1_DelaySelect_Red{7}(2)"
   Button "Button_34" at 595,186 size 38x32; TextOff 'Text'
      on Click: SetTag("DB_HMI_ARG1_Seq1_DelaySelect_Red{8}(2)", 0)
      Visibility <- "DB_HMI_ARG1_Seq1_DelaySelect_Red{8}(2)"
   Button "Button_35" at 665,186 size 38x32; TextOff 'Text'
      on Click: SetTag("DB_HMI_ARG1_Seq1_DelaySelect_Red{9}(2)", 0)
      Visibility <- "DB_HMI_ARG1_Seq1_DelaySelect_Red{9}(2)"
   Button "Button_36" at 735,186 size 38x32; TextOff 'Text'
      on Click: SetTag("DB_HMI_ARG1_Seq1_DelaySelect_Red{10}(2)", 0)
      Visibility <- "DB_HMI_ARG1_Seq1_DelaySelect_Red{10}(2)"
   Button "Button_37" at 176,250 size 38x32; TextOff 'Text'
      on Click: SetTag("DB_HMI_ARG1_Seq1_DelaySelect_Green{2}(2)", 0)
      Visibility <- "DB_HMI_ARG1_Seq1_DelaySelect_Green{2}(2)"
   Button "Button_38" at 246,250 size 38x32; TextOff 'Text'
      on Click: SetTag("DB_HMI_ARG1_Seq1_DelaySelect_Green{3}(2)", 0)
      Visibility <- "DB_HMI_ARG1_Seq1_DelaySelect_Green{3}(2)"
   Button "Button_39" at 316,250 size 38x32; TextOff 'Text'
      on Click: SetTag("DB_HMI_ARG1_Seq1_DelaySelect_Green{4}(2)", 0)
      Visibility <- "DB_HMI_ARG1_Seq1_DelaySelect_Green{4}(2)"
   Button "Button_40" at 386,250 size 38x32; TextOff 'Text'
      on Click: SetTag("DB_HMI_ARG1_Seq1_DelaySelect_Green{5}(2)", 0)
      Visibility <- "DB_HMI_ARG1_Seq1_DelaySelect_Green{5}(2)"
   Button "Button_41" at 456,250 size 38x32; TextOff 'Text'
      on Click: SetTag("DB_HMI_ARG1_Seq1_DelaySelect_Green{6}(2)", 0)
      Visibility <- "DB_HMI_ARG1_Seq1_DelaySelect_Green{6}(2)"
   Button "Button_42" at 526,250 size 38x32; TextOff 'Text'
      on Click: SetTag("DB_HMI_ARG1_Seq1_DelaySelect_Green{7}(2)", 0)
      Visibility <- "DB_HMI_ARG1_Seq1_DelaySelect_Green{7}(2)"
   Button "Button_43" at 596,250 size 38x32; TextOff 'Text'
      on Click: SetTag("DB_HMI_ARG1_Seq1_DelaySelect_Green{8}(2)", 0)
      Visibility <- "DB_HMI_ARG1_Seq1_DelaySelect_Green{8}(2)"
   Button "Button_44" at 666,250 size 38x32; TextOff 'Text'
      on Click: SetTag("DB_HMI_ARG1_Seq1_DelaySelect_Green{9}(2)", 0)
      Visibility <- "DB_HMI_ARG1_Seq1_DelaySelect_Green{9}(2)"
   Button "Button_45" at 736,250 size 38x32; TextOff 'Text'
      on Click: SetTag("DB_HMI_ARG1_Seq1_DelaySelect_Green{10}(2)", 0)
      Visibility <- "DB_HMI_ARG1_Seq1_DelaySelect_Green{10}(2)"
   Button "Button_46" at 176,314 size 38x32; TextOff 'Text'
      on Click: SetTag("DB_HMI_ARG1_Seq1_DelaySelect_Blue{2}(2)", 0)
      Visibility <- "DB_HMI_ARG1_Seq1_DelaySelect_Blue{2}(2)"
   Button "Button_47" at 246,314 size 38x32; TextOff 'Text'
      on Click: SetTag("DB_HMI_ARG1_Seq1_DelaySelect_Blue{3}(2)", 0)
      Visibility <- "DB_HMI_ARG1_Seq1_DelaySelect_Blue{3}(2)"
   Button "Button_48" at 316,314 size 38x32; TextOff 'Text'
      on Click: SetTag("DB_HMI_ARG1_Seq1_DelaySelect_Blue{4}(2)", 0)
      Visibility <- "DB_HMI_ARG1_Seq1_DelaySelect_Blue{4}(2)"
   Button "Button_49" at 386,314 size 38x32; TextOff 'Text'
      on Click: SetTag("DB_HMI_ARG1_Seq1_DelaySelect_Blue{5}(2)", 0)
      Visibility <- "DB_HMI_ARG1_Seq1_DelaySelect_Blue{5}(2)"
   Button "Button_50" at 456,314 size 38x32; TextOff 'Text'
      on Click: SetTag("DB_HMI_ARG1_Seq1_DelaySelect_Blue{6}(2)", 0)
      Visibility <- "DB_HMI_ARG1_Seq1_DelaySelect_Blue{6}(2)"
   Button "Button_51" at 526,314 size 38x32; TextOff 'Text'
      on Click: SetTag("DB_HMI_ARG1_Seq1_DelaySelect_Blue{7}(2)", 0)
      Visibility <- "DB_HMI_ARG1_Seq1_DelaySelect_Blue{7}(2)"
   Button "Button_52" at 596,314 size 38x32; TextOff 'Text'
      on Click: SetTag("DB_HMI_ARG1_Seq1_DelaySelect_Blue{8}(2)", 0)
      Visibility <- "DB_HMI_ARG1_Seq1_DelaySelect_Blue{8}(2)"
   Button "Button_53" at 666,314 size 38x32; TextOff 'Text'
      on Click: SetTag("DB_HMI_ARG1_Seq1_DelaySelect_Blue{9}(2)", 0)
      Visibility <- "DB_HMI_ARG1_Seq1_DelaySelect_Blue{9}(2)"
   Button "Button_54" at 736,314 size 38x32; TextOff 'Text'
      on Click: SetTag("DB_HMI_ARG1_Seq1_DelaySelect_Blue{10}(2)", 0)
      Visibility <- "DB_HMI_ARG1_Seq1_DelaySelect_Blue{10}(2)"
   Button "Button_55" at 619,378 size 165x40; TextOff 'Reset / Alle Quittieren'; PictureOff "More_Icon"
      on ReleaseLeft: ResetBit("Ext_AckSafety_DB_ack")
      on PressLeft: SetBit("Ext_AckSafety_DB_ack")
      on Release: SetTag("DB_HMI_ARG1_Seq1_Cmd_DelayReset(2)", 0)
      on Press: SetTag("DB_HMI_ARG1_Seq1_Cmd_DelayReset(2)", 1)
      ObjectEnable <- "DB_HMI_ARG1_Seq1_Cmd_DelayReset"

screen "40_SimValues_4" 800x480, template "31_SimValues_1"
   GraphicView "gfxDarkBackground" at 0,0 size 800x480; Picture "PopUpBackground"
      Visibility <- "PopUpBackground"
   TextField "txtParameter1_2" at 246,136 size 42x25; Text 'Step 2 / Parameter 1'
   TextField "txtParameter1_3" at 316,136 size 102x25; Text 'Step 3 / Parameter 1'
   TextField "txtParameter1_4" at 386,136 size 102x25; Text 'Step 4 / Parameter 1'
   TextField "txtParameter1_5" at 456,136 size 102x25; Text 'Step 5 / Parameter 1'
   TextField "txtParameter1_6" at 526,136 size 102x25; Text 'Step 6 / Parameter 1'
   TextField "txtParameter1_8" at 596,136 size 102x25; Text 'Step 7 / Parameter 1'
   TextField "txtParameter1_9" at 666,136 size 102x25; Text 'Step 8 / Parameter 1'
   TextField "txtParameter1_10" at 176,136 size 45x25; Text 'Step 1 / Parameter 1'
   TextField "txtParameter1_11" at 736,136 size 46x25; Text 'Step 9 / Parameter 1'
   TextField "txtParameter1_1" at 104,136 size 45x25; Text 'Branch / Parameter 1'
   TextField "txtParameter1_7" at 32,136 size 45x25; Text 'Car / Parameter 1'
   GraphicView "Graphic view_1" at 33,184 size 40x40; Picture "Car_Red"
   GraphicView "Graphic view_3" at 33,249 size 40x40; Picture "Car_Green"
   GraphicView "Graphic view_4" at 33,308 size 40x40; Picture "Car_Blue_1"
   TextField "Text field_3" at 121,191 size 15x23; Text '1'
      Visibility <- "InScreenTabState"
   TextField "Text field_1" at 121,256 size 15x23; Text '2'
      Visibility <- "InScreenTabState"
   TextField "Text field_2" at 121,321 size 15x23; Text '2'
      Visibility <- "InScreenTabState"
   Button "Button_1" at 176,186 size 38x32; TextOff 'Text'
      on Click: SetTag("DB_HMI_ARG1_Seq1_DelaySelect_Red{2}(3)", 1)
   Button "Button_2" at 245,186 size 38x32; TextOff 'Text'
      on Click: SetTag("DB_HMI_ARG1_Seq1_DelaySelect_Red{3}(3)", 1)
   Button "Button_3" at 315,186 size 38x32; TextOff 'Text'
      on Click: SetTag("DB_HMI_ARG1_Seq1_DelaySelect_Red{4}(3)", 1)
   Button "Button_4" at 385,186 size 38x32; TextOff 'Text'
      on Click: SetTag("DB_HMI_ARG1_Seq1_DelaySelect_Red{5}(3)", 1)
   Button "Button_5" at 455,186 size 38x32; TextOff 'Text'
      on Click: SetTag("DB_HMI_ARG1_Seq1_DelaySelect_Red{6}(3)", 1)
   Button "Button_6" at 525,186 size 38x32; TextOff 'Text'
      on Click: SetTag("DB_HMI_ARG1_Seq1_DelaySelect_Red{7}(3)", 1)
   Button "Button_8" at 595,186 size 38x32; TextOff 'Text'
      on Click: SetTag("DB_HMI_ARG1_Seq1_DelaySelect_Red{8}(3)", 1)
   Button "Button_9" at 665,186 size 38x32; TextOff 'Text'
      on Click: SetTag("DB_HMI_ARG1_Seq1_DelaySelect_Red{9}(3)", 1)
   Button "Button_10" at 735,186 size 38x32; TextOff 'Text'
      on Click: SetTag("DB_HMI_ARG1_Seq1_DelaySelect_Red{10}(3)", 1)
   Button "Button_17" at 176,250 size 38x32; TextOff 'Text'
      on Click: SetTag("DB_HMI_ARG1_Seq1_DelaySelect_Green{2}(3)", 1)
   Button "Button_7" at 246,250 size 38x32; TextOff 'Text'
      on Click: SetTag("DB_HMI_ARG1_Seq1_DelaySelect_Green{3}(3)", 1)
   Button "Button_11" at 316,250 size 38x32; TextOff 'Text'
      on Click: SetTag("DB_HMI_ARG1_Seq1_DelaySelect_Green{4}(3)", 1)
   Button "Button_12" at 386,250 size 38x32; TextOff 'Text'
      on Click: SetTag("DB_HMI_ARG1_Seq1_DelaySelect_Green{5}(3)", 1)
   Button "Button_13" at 456,250 size 38x32; TextOff 'Text'
      on Click: SetTag("DB_HMI_ARG1_Seq1_DelaySelect_Green{6}(3)", 1)
   Button "Button_14" at 526,250 size 38x32; TextOff 'Text'
      on Click: SetTag("DB_HMI_ARG1_Seq1_DelaySelect_Green{7}(3)", 1)
   Button "Button_15" at 596,250 size 38x32; TextOff 'Text'
      on Click: SetTag("DB_HMI_ARG1_Seq1_DelaySelect_Green{8}(3)", 1)
   Button "Button_16" at 666,250 size 38x32; TextOff 'Text'
      on Click: SetTag("DB_HMI_ARG1_Seq1_DelaySelect_Green{9}(3)", 1)
   Button "Button_18" at 736,250 size 38x32; TextOff 'Text'
      on Click: SetTag("DB_HMI_ARG1_Seq1_DelaySelect_Green{10}(3)", 1)
   Button "Button_26" at 176,314 size 38x32; TextOff 'Text'
      on Click: SetTag("DB_HMI_ARG1_Seq1_DelaySelect_Blue{2}(3)", 1)
   Button "Button_19" at 246,314 size 38x32; TextOff 'Text'
      on Click: SetTag("DB_HMI_ARG1_Seq1_DelaySelect_Blue{3}(3)", 1)
   Button "Button_20" at 316,314 size 38x32; TextOff 'Text'
      on Click: SetTag("DB_HMI_ARG1_Seq1_DelaySelect_Blue{4}(3)", 1)
   Button "Button_21" at 386,314 size 38x32; TextOff 'Text'
      on Click: SetTag("DB_HMI_ARG1_Seq1_DelaySelect_Blue{5}(3)", 1)
   Button "Button_22" at 456,314 size 38x32; TextOff 'Text'
      on Click: SetTag("DB_HMI_ARG1_Seq1_DelaySelect_Blue{6}(3)", 1)
   Button "Button_23" at 526,314 size 38x32; TextOff 'Text'
      on Click: SetTag("DB_HMI_ARG1_Seq1_DelaySelect_Blue{7}(3)", 1)
   Button "Button_24" at 596,314 size 38x32; TextOff 'Text'
      on Click: SetTag("DB_HMI_ARG1_Seq1_DelaySelect_Blue{8}(3)", 1)
   Button "Button_25" at 666,314 size 38x32; TextOff 'Text'
      on Click: SetTag("DB_HMI_ARG1_Seq1_DelaySelect_Blue{9}(3)", 1)
   Button "Button_27" at 736,314 size 38x32; TextOff 'Text'
      on Click: SetTag("DB_HMI_ARG1_Seq1_DelaySelect_Blue{10}(3)", 1)
   Button "Button_28" at 176,186 size 38x32; TextOff 'Text'
      on Click: SetTag("DB_HMI_ARG1_Seq1_DelaySelect_Red{2}(3)", 0)
      Visibility <- "DB_HMI_ARG1_Seq1_DelaySelect_Red{2}(3)"
   Button "Button_29" at 245,186 size 38x32; TextOff 'Text'
      on Click: SetTag("DB_HMI_ARG1_Seq1_DelaySelect_Red{3}(3)", 0)
      Visibility <- "DB_HMI_ARG1_Seq1_DelaySelect_Red{3}(3)"
   Button "Button_30" at 315,186 size 38x32; TextOff 'Text'
      on Click: SetTag("DB_HMI_ARG1_Seq1_DelaySelect_Red{4}(3)", 0)
      Visibility <- "DB_HMI_ARG1_Seq1_DelaySelect_Red{4}(3)"
   Button "Button_31" at 385,186 size 38x32; TextOff 'Text'
      on Click: SetTag("DB_HMI_ARG1_Seq1_DelaySelect_Red{5}(3)", 0)
      Visibility <- "DB_HMI_ARG1_Seq1_DelaySelect_Red{5}(3)"
   Button "Button_32" at 455,186 size 38x32; TextOff 'Text'
      on Click: SetTag("DB_HMI_ARG1_Seq1_DelaySelect_Red{6}(3)", 0)
      Visibility <- "DB_HMI_ARG1_Seq1_DelaySelect_Red{6}(3)"
   Button "Button_33" at 525,186 size 38x32; TextOff 'Text'
      on Click: SetTag("DB_HMI_ARG1_Seq1_DelaySelect_Red{7}(3)", 0)
      Visibility <- "DB_HMI_ARG1_Seq1_DelaySelect_Red{7}(3)"
   Button "Button_34" at 595,186 size 38x32; TextOff 'Text'
      on Click: SetTag("DB_HMI_ARG1_Seq1_DelaySelect_Red{8}(3)", 0)
      Visibility <- "DB_HMI_ARG1_Seq1_DelaySelect_Red{8}(3)"
   Button "Button_35" at 665,186 size 38x32; TextOff 'Text'
      on Click: SetTag("DB_HMI_ARG1_Seq1_DelaySelect_Red{9}(3)", 0)
      Visibility <- "DB_HMI_ARG1_Seq1_DelaySelect_Red{9}(3)"
   Button "Button_36" at 735,186 size 38x32; TextOff 'Text'
      on Click: SetTag("DB_HMI_ARG1_Seq1_DelaySelect_Red{10}(3)", 0)
      Visibility <- "DB_HMI_ARG1_Seq1_DelaySelect_Red{10}(3)"
   Button "Button_37" at 176,250 size 38x32; TextOff 'Text'
      on Click: SetTag("DB_HMI_ARG1_Seq1_DelaySelect_Green{2}(3)", 0)
      Visibility <- "DB_HMI_ARG1_Seq1_DelaySelect_Green{2}(3)"
   Button "Button_38" at 246,250 size 38x32; TextOff 'Text'
      on Click: SetTag("DB_HMI_ARG1_Seq1_DelaySelect_Green{3}(3)", 0)
      Visibility <- "DB_HMI_ARG1_Seq1_DelaySelect_Green{3}(3)"
   Button "Button_39" at 316,250 size 38x32; TextOff 'Text'
      on Click: SetTag("DB_HMI_ARG1_Seq1_DelaySelect_Green{4}(3)", 0)
      Visibility <- "DB_HMI_ARG1_Seq1_DelaySelect_Green{4}(3)"
   Button "Button_40" at 386,250 size 38x32; TextOff 'Text'
      on Click: SetTag("DB_HMI_ARG1_Seq1_DelaySelect_Green{5}(3)", 0)
      Visibility <- "DB_HMI_ARG1_Seq1_DelaySelect_Green{5}(3)"
   Button "Button_41" at 456,250 size 38x32; TextOff 'Text'
      on Click: SetTag("DB_HMI_ARG1_Seq1_DelaySelect_Green{6}(3)", 0)
      Visibility <- "DB_HMI_ARG1_Seq1_DelaySelect_Green{6}(3)"
   Button "Button_42" at 526,250 size 38x32; TextOff 'Text'
      on Click: SetTag("DB_HMI_ARG1_Seq1_DelaySelect_Green{7}(3)", 0)
      Visibility <- "DB_HMI_ARG1_Seq1_DelaySelect_Green{7}(3)"
   Button "Button_43" at 596,250 size 38x32; TextOff 'Text'
      on Click: SetTag("DB_HMI_ARG1_Seq1_DelaySelect_Green{8}(3)", 0)
      Visibility <- "DB_HMI_ARG1_Seq1_DelaySelect_Green{8}(3)"
   Button "Button_44" at 666,250 size 38x32; TextOff 'Text'
      on Click: SetTag("DB_HMI_ARG1_Seq1_DelaySelect_Green{9}(3)", 0)
      Visibility <- "DB_HMI_ARG1_Seq1_DelaySelect_Green{9}(3)"
   Button "Button_45" at 736,250 size 38x32; TextOff 'Text'
      on Click: SetTag("DB_HMI_ARG1_Seq1_DelaySelect_Green{10}(3)", 0)
      Visibility <- "DB_HMI_ARG1_Seq1_DelaySelect_Green{10}(3)"
   Button "Button_46" at 176,314 size 38x32; TextOff 'Text'
      on Click: SetTag("DB_HMI_ARG1_Seq1_DelaySelect_Blue{2}(3)", 0)
      Visibility <- "DB_HMI_ARG1_Seq1_DelaySelect_Blue{2}(3)"
   Button "Button_47" at 246,314 size 38x32; TextOff 'Text'
      on Click: SetTag("DB_HMI_ARG1_Seq1_DelaySelect_Blue{3}(3)", 0)
      Visibility <- "DB_HMI_ARG1_Seq1_DelaySelect_Blue{3}(3)"
   Button "Button_48" at 316,314 size 38x32; TextOff 'Text'
      on Click: SetTag("DB_HMI_ARG1_Seq1_DelaySelect_Blue{4}(3)", 0)
      Visibility <- "DB_HMI_ARG1_Seq1_DelaySelect_Blue{4}(3)"
   Button "Button_49" at 386,314 size 38x32; TextOff 'Text'
      on Click: SetTag("DB_HMI_ARG1_Seq1_DelaySelect_Blue{5}(3)", 0)
      Visibility <- "DB_HMI_ARG1_Seq1_DelaySelect_Blue{5}(3)"
   Button "Button_50" at 456,314 size 38x32; TextOff 'Text'
      on Click: SetTag("DB_HMI_ARG1_Seq1_DelaySelect_Blue{6}(3)", 0)
      Visibility <- "DB_HMI_ARG1_Seq1_DelaySelect_Blue{6}(3)"
   Button "Button_51" at 526,314 size 38x32; TextOff 'Text'
      on Click: SetTag("DB_HMI_ARG1_Seq1_DelaySelect_Blue{7}(3)", 0)
      Visibility <- "DB_HMI_ARG1_Seq1_DelaySelect_Blue{7}(3)"
   Button "Button_52" at 596,314 size 38x32; TextOff 'Text'
      on Click: SetTag("DB_HMI_ARG1_Seq1_DelaySelect_Blue{8}(3)", 0)
      Visibility <- "DB_HMI_ARG1_Seq1_DelaySelect_Blue{8}(3)"
   Button "Button_53" at 666,314 size 38x32; TextOff 'Text'
      on Click: SetTag("DB_HMI_ARG1_Seq1_DelaySelect_Blue{9}(3)", 0)
      Visibility <- "DB_HMI_ARG1_Seq1_DelaySelect_Blue{9}(3)"
   Button "Button_54" at 736,314 size 38x32; TextOff 'Text'
      on Click: SetTag("DB_HMI_ARG1_Seq1_DelaySelect_Blue{10}(3)", 0)
      Visibility <- "DB_HMI_ARG1_Seq1_DelaySelect_Blue{10}(3)"
   Button "Button_55" at 619,378 size 165x40; TextOff 'Reset / Alle Quittieren'; PictureOff "More_Icon"
      on ReleaseLeft: ResetBit("Ext_AckSafety_DB_ack")
      on PressLeft: SetBit("Ext_AckSafety_DB_ack")
      on Release: SetTag("DB_HMI_ARG1_Seq1_Cmd_DelayReset(3)", 0)
      on Press: SetTag("DB_HMI_ARG1_Seq1_Cmd_DelayReset(3)", 1)
      ObjectEnable <- "DB_HMI_ARG1_Seq1_Cmd_DelayReset"

